   
   	SmartTags("SDC\DB_SDC_ERROR_STAT\_Byte_DB_SDC_ERROR_STAT.F_STAT[XX1].EMS_TS_STAT_VAL.PROFIL") =  			  2 + Eintrag_0 * Laenge_FAULT - Laenge_FAULT + Allg_Offset
   	SmartTags("SDC\DB_SDC_ERROR_STAT\_Byte_DB_SDC_ERROR_STAT.F_STAT[XX2].EMS_TS_STAT_VAL.PROFIL") =  			  2 + Eintrag_1 * Laenge_FAULT - Laenge_FAULT + Allg_Offset
   	SmartTags("SDC\DB_SDC_ERROR_STAT\_Byte_DB_SDC_ERROR_STAT.F_STAT[XX3].EMS_TS_STAT_VAL.PROFIL") =  			  2 + Eintrag_2 * Laenge_FAULT - Laenge_FAULT + Allg_Offset
   	SmartTags("SDC\DB_SDC_ERROR_STAT\_Byte_DB_SDC_ERROR_STAT.F_STAT[XX4].EMS_TS_STAT_VAL.PROFIL") =  			  2 + Eintrag_3 * Laenge_FAULT - Laenge_FAULT + Allg_Offset
   	SmartTags("SDC\DB_SDC_ERROR_STAT\_Byte_DB_SDC_ERROR_STAT.F_STAT[XX5].EMS_TS_STAT_VAL.PROFIL") =  			  2 + Eintrag_4 * Laenge_FAULT - Laenge_FAULT + Allg_Offset
   	SmartTags("SDC\DB_SDC_ERROR_STAT\_Byte_DB_SDC_ERROR_STAT.F_STAT[XX6].EMS_TS_STAT_VAL.PROFIL") =  			  2 + Eintrag_5 * Laenge_FAULT - Laenge_FAULT + Allg_Offset
   	SmartTags("SDC\DB_SDC_ERROR_STAT\_Byte_DB_SDC_ERROR_STAT.F_STAT[XX7].EMS_TS_STAT_VAL.PROFIL") =  			  2 + Eintrag_6 * Laenge_FAULT - Laenge_FAULT + Allg_Offset
   	SmartTags("SDC\DB_SDC_ERROR_STAT\_Byte_DB_SDC_ERROR_STAT.F_STAT[XX8].EMS_TS_STAT_VAL.PROFIL") =  			  2 + Eintrag_7 * Laenge_FAULT - Laenge_FAULT + Allg_Offset
   	SmartTags("SDC\DB_SDC_ERROR_STAT\_Byte_DB_SDC_ERROR_STAT.F_STAT[XX9].EMS_TS_STAT_VAL.PROFIL") =  			  2 + Eintrag_8 * Laenge_FAULT - Laenge_FAULT + Allg_Offset
   	SmartTags("SDC\DB_SDC_ERROR_STAT\_Byte_DB_SDC_ERROR_STAT.F_STAT[X10].EMS_TS_STAT_VAL.PROFIL") =  			  2 + Eintrag_9 * Laenge_FAULT - Laenge_FAULT + Allg_Offset
   
   	SmartTags("SDC\DB_SDC_ERROR_STAT\_Byte_DB_SDC_ERROR_STAT.F_STAT[XX1].EMS_TS_STAT_VAL.DRIVE_POS") =   		  4 + Eintrag_0 * Laenge_FAULT - Laenge_FAULT + Allg_Offset
   	SmartTags("SDC\DB_SDC_ERROR_STAT\_Byte_DB_SDC_ERROR_STAT.F_STAT[XX2].EMS_TS_STAT_VAL.DRIVE_POS") =   		  4 + Eintrag_1 * Laenge_FAULT - Laenge_FAULT + Allg_Offset
   	SmartTags("SDC\DB_SDC_ERROR_STAT\_Byte_DB_SDC_ERROR_STAT.F_STAT[XX3].EMS_TS_STAT_VAL.DRIVE_POS") =   		  4 + Eintrag_2 * Laenge_FAULT - Laenge_FAULT + Allg_Offset
   	SmartTags("SDC\DB_SDC_ERROR_STAT\_Byte_DB_SDC_ERROR_STAT.F_STAT[XX4].EMS_TS_STAT_VAL.DRIVE_POS") =   		  4 + Eintrag_3 * Laenge_FAULT - Laenge_FAULT + Allg_Offset
   	SmartTags("SDC\DB_SDC_ERROR_STAT\_Byte_DB_SDC_ERROR_STAT.F_STAT[XX5].EMS_TS_STAT_VAL.DRIVE_POS") =   		  4 + Eintrag_4 * Laenge_FAULT - Laenge_FAULT + Allg_Offset
   	SmartTags("SDC\DB_SDC_ERROR_STAT\_Byte_DB_SDC_ERROR_STAT.F_STAT[XX6].EMS_TS_STAT_VAL.DRIVE_POS") =   		  4 + Eintrag_5 * Laenge_FAULT - Laenge_FAULT + Allg_Offset
   	SmartTags("SDC\DB_SDC_ERROR_STAT\_Byte_DB_SDC_ERROR_STAT.F_STAT[XX7].EMS_TS_STAT_VAL.DRIVE_POS") =   		  4 + Eintrag_6 * Laenge_FAULT - Laenge_FAULT + Allg_Offset
   	SmartTags("SDC\DB_SDC_ERROR_STAT\_Byte_DB_SDC_ERROR_STAT.F_STAT[XX8].EMS_TS_STAT_VAL.DRIVE_POS") =   		  4 + Eintrag_7 * Laenge_FAULT - Laenge_FAULT + Allg_Offset
   	SmartTags("SDC\DB_SDC_ERROR_STAT\_Byte_DB_SDC_ERROR_STAT.F_STAT[XX9].EMS_TS_STAT_VAL.DRIVE_POS") =   		  4 + Eintrag_8 * Laenge_FAULT - Laenge_FAULT + Allg_Offset
   	SmartTags("SDC\DB_SDC_ERROR_STAT\_Byte_DB_SDC_ERROR_STAT.F_STAT[X10].EMS_TS_STAT_VAL.DRIVE_POS") =   		  4 + Eintrag_9 * Laenge_FAULT - Laenge_FAULT + Allg_Offset
   	
   	SmartTags("SDC\DB_SDC_ERROR_STAT\_Byte_DB_SDC_ERROR_STAT.F_STAT[XX1].EMS_TS_STAT_VAL.HOIST_POS") =   		  8 + Eintrag_0 * Laenge_FAULT - Laenge_FAULT + Allg_Offset
   	SmartTags("SDC\DB_SDC_ERROR_STAT\_Byte_DB_SDC_ERROR_STAT.F_STAT[XX2].EMS_TS_STAT_VAL.HOIST_POS") =   		  8 + Eintrag_1 * Laenge_FAULT - Laenge_FAULT + Allg_Offset
   	SmartTags("SDC\DB_SDC_ERROR_STAT\_Byte_DB_SDC_ERROR_STAT.F_STAT[XX3].EMS_TS_STAT_VAL.HOIST_POS") =   		  8 + Eintrag_2 * Laenge_FAULT - Laenge_FAULT + Allg_Offset
   	SmartTags("SDC\DB_SDC_ERROR_STAT\_Byte_DB_SDC_ERROR_STAT.F_STAT[XX4].EMS_TS_STAT_VAL.HOIST_POS") =   		  8 + Eintrag_3 * Laenge_FAULT - Laenge_FAULT + Allg_Offset
   	SmartTags("SDC\DB_SDC_ERROR_STAT\_Byte_DB_SDC_ERROR_STAT.F_STAT[XX5].EMS_TS_STAT_VAL.HOIST_POS") =   		  8 + Eintrag_4 * Laenge_FAULT - Laenge_FAULT + Allg_Offset
   	SmartTags("SDC\DB_SDC_ERROR_STAT\_Byte_DB_SDC_ERROR_STAT.F_STAT[XX6].EMS_TS_STAT_VAL.HOIST_POS") =   		  8 + Eintrag_5 * Laenge_FAULT - Laenge_FAULT + Allg_Offset
   	SmartTags("SDC\DB_SDC_ERROR_STAT\_Byte_DB_SDC_ERROR_STAT.F_STAT[XX7].EMS_TS_STAT_VAL.HOIST_POS") =   		  8 + Eintrag_6 * Laenge_FAULT - Laenge_FAULT + Allg_Offset
   	SmartTags("SDC\DB_SDC_ERROR_STAT\_Byte_DB_SDC_ERROR_STAT.F_STAT[XX8].EMS_TS_STAT_VAL.HOIST_POS") =   		  8 + Eintrag_7 * Laenge_FAULT - Laenge_FAULT + Allg_Offset
   	SmartTags("SDC\DB_SDC_ERROR_STAT\_Byte_DB_SDC_ERROR_STAT.F_STAT[XX9].EMS_TS_STAT_VAL.HOIST_POS") =   		  8 + Eintrag_8 * Laenge_FAULT - Laenge_FAULT + Allg_Offset
   	SmartTags("SDC\DB_SDC_ERROR_STAT\_Byte_DB_SDC_ERROR_STAT.F_STAT[X10].EMS_TS_STAT_VAL.HOIST_POS") =   		  8 + Eintrag_9 * Laenge_FAULT - Laenge_FAULT + Allg_Offset
   	
   '	SmartTags("SDC\DB_SDC_ERROR_STAT\_Byte_DB_SDC_ERROR_STAT.F_STAT[XX1].EMS_TS_STAT_VAL.TILT_POS")  =   		 10 + Eintrag_0 * Laenge_FAULT - Laenge_FAULT + Allg_Offset
   '	SmartTags("SDC\DB_SDC_ERROR_STAT\_Byte_DB_SDC_ERROR_STAT.F_STAT[XX2].EMS_TS_STAT_VAL.TILT_POS")  =   		 10 + Eintrag_1 * Laenge_FAULT - Laenge_FAULT + Allg_Offset
   '	SmartTags("SDC\DB_SDC_ERROR_STAT\_Byte_DB_SDC_ERROR_STAT.F_STAT[XX3].EMS_TS_STAT_VAL.TILT_POS")  =   		 10 + Eintrag_2 * Laenge_FAULT - Laenge_FAULT + Allg_Offset
   '	SmartTags("SDC\DB_SDC_ERROR_STAT\_Byte_DB_SDC_ERROR_STAT.F_STAT[XX4].EMS_TS_STAT_VAL.TILT_POS")  =   		 10 + Eintrag_3 * Laenge_FAULT - Laenge_FAULT + Allg_Offset
   '	SmartTags("SDC\DB_SDC_ERROR_STAT\_Byte_DB_SDC_ERROR_STAT.F_STAT[XX5].EMS_TS_STAT_VAL.TILT_POS")  =   		 10 + Eintrag_4 * Laenge_FAULT - Laenge_FAULT + Allg_Offset
   '	SmartTags("SDC\DB_SDC_ERROR_STAT\_Byte_DB_SDC_ERROR_STAT.F_STAT[XX6].EMS_TS_STAT_VAL.TILT_POS")  =   		 10 + Eintrag_5 * Laenge_FAULT - Laenge_FAULT + Allg_Offset
   '	SmartTags("SDC\DB_SDC_ERROR_STAT\_Byte_DB_SDC_ERROR_STAT.F_STAT[XX7].EMS_TS_STAT_VAL.TILT_POS")  =   		 10 + Eintrag_6 * Laenge_FAULT - Laenge_FAULT + Allg_Offset
   '	SmartTags("SDC\DB_SDC_ERROR_STAT\_Byte_DB_SDC_ERROR_STAT.F_STAT[XX8].EMS_TS_STAT_VAL.TILT_POS")  =   		 10 + Eintrag_7 * Laenge_FAULT - Laenge_FAULT + Allg_Offset
   '	SmartTags("SDC\DB_SDC_ERROR_STAT\_Byte_DB_SDC_ERROR_STAT.F_STAT[XX9].EMS_TS_STAT_VAL.TILT_POS")  =   		 10 + Eintrag_8 * Laenge_FAULT - Laenge_FAULT + Allg_Offset
   '	SmartTags("SDC\DB_SDC_ERROR_STAT\_Byte_DB_SDC_ERROR_STAT.F_STAT[X10].EMS_TS_STAT_VAL.TILT_POS")  =   		 10 + Eintrag_9 * Laenge_FAULT - Laenge_FAULT + Allg_Offset
   	
   	SmartTags("SDC\DB_SDC_ERROR_STAT\_Byte_DB_SDC_ERROR_STAT.F_STAT[XX1].EMS_TS_STAT_VAL.ERROR")  	 =   		 10 + Eintrag_0 * Laenge_FAULT - Laenge_FAULT + Allg_Offset
   	SmartTags("SDC\DB_SDC_ERROR_STAT\_Byte_DB_SDC_ERROR_STAT.F_STAT[XX2].EMS_TS_STAT_VAL.ERROR")  	 =   		 10 + Eintrag_1 * Laenge_FAULT - Laenge_FAULT + Allg_Offset
   	SmartTags("SDC\DB_SDC_ERROR_STAT\_Byte_DB_SDC_ERROR_STAT.F_STAT[XX3].EMS_TS_STAT_VAL.ERROR")  	 =   		 10 + Eintrag_2 * Laenge_FAULT - Laenge_FAULT + Allg_Offset
   	SmartTags("SDC\DB_SDC_ERROR_STAT\_Byte_DB_SDC_ERROR_STAT.F_STAT[XX4].EMS_TS_STAT_VAL.ERROR")  	 =   		 10 + Eintrag_3 * Laenge_FAULT - Laenge_FAULT + Allg_Offset
   	SmartTags("SDC\DB_SDC_ERROR_STAT\_Byte_DB_SDC_ERROR_STAT.F_STAT[XX5].EMS_TS_STAT_VAL.ERROR")  	 =   		 10 + Eintrag_4 * Laenge_FAULT - Laenge_FAULT + Allg_Offset
   	SmartTags("SDC\DB_SDC_ERROR_STAT\_Byte_DB_SDC_ERROR_STAT.F_STAT[XX6].EMS_TS_STAT_VAL.ERROR")  	 =   		 10 + Eintrag_5 * Laenge_FAULT - Laenge_FAULT + Allg_Offset
   	SmartTags("SDC\DB_SDC_ERROR_STAT\_Byte_DB_SDC_ERROR_STAT.F_STAT[XX7].EMS_TS_STAT_VAL.ERROR")  	 =   		 10 + Eintrag_6 * Laenge_FAULT - Laenge_FAULT + Allg_Offset
   	SmartTags("SDC\DB_SDC_ERROR_STAT\_Byte_DB_SDC_ERROR_STAT.F_STAT[XX8].EMS_TS_STAT_VAL.ERROR")  	 =   		 10 + Eintrag_7 * Laenge_FAULT - Laenge_FAULT + Allg_Offset
   	SmartTags("SDC\DB_SDC_ERROR_STAT\_Byte_DB_SDC_ERROR_STAT.F_STAT[XX9].EMS_TS_STAT_VAL.ERROR")  	 =   		 10 + Eintrag_8 * Laenge_FAULT - Laenge_FAULT + Allg_Offset
   	SmartTags("SDC\DB_SDC_ERROR_STAT\_Byte_DB_SDC_ERROR_STAT.F_STAT[X10].EMS_TS_STAT_VAL.ERROR")  	 =   		 10 + Eintrag_9 * Laenge_FAULT - Laenge_FAULT + Allg_Offset
   
   	SmartTags("SDC\DB_SDC_ERROR_STAT\_Byte_DB_SDC_ERROR_STAT.F_STAT[XX1].EMS_TS_STAT_VAL.DRIVE_POS_PERC") =   	 12 + Eintrag_0 * Laenge_FAULT - Laenge_FAULT + Allg_Offset
   	SmartTags("SDC\DB_SDC_ERROR_STAT\_Byte_DB_SDC_ERROR_STAT.F_STAT[XX2].EMS_TS_STAT_VAL.DRIVE_POS_PERC") =   	 12 + Eintrag_1 * Laenge_FAULT - Laenge_FAULT + Allg_Offset
   	SmartTags("SDC\DB_SDC_ERROR_STAT\_Byte_DB_SDC_ERROR_STAT.F_STAT[XX3].EMS_TS_STAT_VAL.DRIVE_POS_PERC") =   	 12 + Eintrag_2 * Laenge_FAULT - Laenge_FAULT + Allg_Offset
   	SmartTags("SDC\DB_SDC_ERROR_STAT\_Byte_DB_SDC_ERROR_STAT.F_STAT[XX4].EMS_TS_STAT_VAL.DRIVE_POS_PERC") =   	 12 + Eintrag_3 * Laenge_FAULT - Laenge_FAULT + Allg_Offset
   	SmartTags("SDC\DB_SDC_ERROR_STAT\_Byte_DB_SDC_ERROR_STAT.F_STAT[XX5].EMS_TS_STAT_VAL.DRIVE_POS_PERC") =   	 12 + Eintrag_4 * Laenge_FAULT - Laenge_FAULT + Allg_Offset
   	SmartTags("SDC\DB_SDC_ERROR_STAT\_Byte_DB_SDC_ERROR_STAT.F_STAT[XX6].EMS_TS_STAT_VAL.DRIVE_POS_PERC") =   	 12 + Eintrag_5 * Laenge_FAULT - Laenge_FAULT + Allg_Offset
   	SmartTags("SDC\DB_SDC_ERROR_STAT\_Byte_DB_SDC_ERROR_STAT.F_STAT[XX7].EMS_TS_STAT_VAL.DRIVE_POS_PERC") =   	 12 + Eintrag_6 * Laenge_FAULT - Laenge_FAULT + Allg_Offset
   	SmartTags("SDC\DB_SDC_ERROR_STAT\_Byte_DB_SDC_ERROR_STAT.F_STAT[XX8].EMS_TS_STAT_VAL.DRIVE_POS_PERC") =   	 12 + Eintrag_7 * Laenge_FAULT - Laenge_FAULT + Allg_Offset
   	SmartTags("SDC\DB_SDC_ERROR_STAT\_Byte_DB_SDC_ERROR_STAT.F_STAT[XX9].EMS_TS_STAT_VAL.DRIVE_POS_PERC") =   	 12 + Eintrag_8 * Laenge_FAULT - Laenge_FAULT + Allg_Offset
   	SmartTags("SDC\DB_SDC_ERROR_STAT\_Byte_DB_SDC_ERROR_STAT.F_STAT[X10].EMS_TS_STAT_VAL.DRIVE_POS_PERC") =   	 12 + Eintrag_9 * Laenge_FAULT - Laenge_FAULT + Allg_Offset
   	
   	SmartTags("SDC\DB_SDC_ERROR_STAT\_Byte_DB_SDC_ERROR_STAT.F_STAT[XX1].EMS_TS_STAT_VAL.SEK") 			=   	 14 + Eintrag_0 * Laenge_FAULT - Laenge_FAULT + Allg_Offset
   	SmartTags("SDC\DB_SDC_ERROR_STAT\_Byte_DB_SDC_ERROR_STAT.F_STAT[XX2].EMS_TS_STAT_VAL.SEK") 			=   	 14 + Eintrag_1 * Laenge_FAULT - Laenge_FAULT + Allg_Offset
   	SmartTags("SDC\DB_SDC_ERROR_STAT\_Byte_DB_SDC_ERROR_STAT.F_STAT[XX3].EMS_TS_STAT_VAL.SEK") 			=   	 14 + Eintrag_2 * Laenge_FAULT - Laenge_FAULT + Allg_Offset
   	SmartTags("SDC\DB_SDC_ERROR_STAT\_Byte_DB_SDC_ERROR_STAT.F_STAT[XX4].EMS_TS_STAT_VAL.SEK") 			=   	 14 + Eintrag_3 * Laenge_FAULT - Laenge_FAULT + Allg_Offset
   	SmartTags("SDC\DB_SDC_ERROR_STAT\_Byte_DB_SDC_ERROR_STAT.F_STAT[XX5].EMS_TS_STAT_VAL.SEK") 			=   	 14 + Eintrag_4 * Laenge_FAULT - Laenge_FAULT + Allg_Offset
   	SmartTags("SDC\DB_SDC_ERROR_STAT\_Byte_DB_SDC_ERROR_STAT.F_STAT[XX6].EMS_TS_STAT_VAL.SEK") 			=   	 14 + Eintrag_5 * Laenge_FAULT - Laenge_FAULT + Allg_Offset
   	SmartTags("SDC\DB_SDC_ERROR_STAT\_Byte_DB_SDC_ERROR_STAT.F_STAT[XX7].EMS_TS_STAT_VAL.SEK") 			=   	 14 + Eintrag_6 * Laenge_FAULT - Laenge_FAULT + Allg_Offset
   	SmartTags("SDC\DB_SDC_ERROR_STAT\_Byte_DB_SDC_ERROR_STAT.F_STAT[XX8].EMS_TS_STAT_VAL.SEK") 			=   	 14 + Eintrag_7 * Laenge_FAULT - Laenge_FAULT + Allg_Offset
   	SmartTags("SDC\DB_SDC_ERROR_STAT\_Byte_DB_SDC_ERROR_STAT.F_STAT[XX9].EMS_TS_STAT_VAL.SEK") 			=   	 14 + Eintrag_8 * Laenge_FAULT - Laenge_FAULT + Allg_Offset
   	SmartTags("SDC\DB_SDC_ERROR_STAT\_Byte_DB_SDC_ERROR_STAT.F_STAT[X10].EMS_TS_STAT_VAL.SEK") 			=   	 14 + Eintrag_9 * Laenge_FAULT - Laenge_FAULT + Allg_Offset
   	
   	SmartTags("SDC\DB_SDC_ERROR_STAT\_Byte_DB_SDC_ERROR_STAT.F_STAT[XX1].F") = 									 16 + Eintrag_0 * Laenge_FAULT - Laenge_FAULT + Allg_Offset
   	SmartTags("SDC\DB_SDC_ERROR_STAT\_Byte_DB_SDC_ERROR_STAT.F_STAT[XX2].F") = 									 16 + Eintrag_1 * Laenge_FAULT - Laenge_FAULT + Allg_Offset
   	SmartTags("SDC\DB_SDC_ERROR_STAT\_Byte_DB_SDC_ERROR_STAT.F_STAT[XX3].F") = 									 16 + Eintrag_2 * Laenge_FAULT - Laenge_FAULT + Allg_Offset
   	SmartTags("SDC\DB_SDC_ERROR_STAT\_Byte_DB_SDC_ERROR_STAT.F_STAT[XX4].F") = 									 16 + Eintrag_3 * Laenge_FAULT - Laenge_FAULT + Allg_Offset
   	SmartTags("SDC\DB_SDC_ERROR_STAT\_Byte_DB_SDC_ERROR_STAT.F_STAT[XX5].F") = 									 16 + Eintrag_4 * Laenge_FAULT - Laenge_FAULT + Allg_Offset
   	SmartTags("SDC\DB_SDC_ERROR_STAT\_Byte_DB_SDC_ERROR_STAT.F_STAT[XX6].F") = 									 16 + Eintrag_5 * Laenge_FAULT - Laenge_FAULT + Allg_Offset
   	SmartTags("SDC\DB_SDC_ERROR_STAT\_Byte_DB_SDC_ERROR_STAT.F_STAT[XX7].F") = 									 16 + Eintrag_6 * Laenge_FAULT - Laenge_FAULT + Allg_Offset
   	SmartTags("SDC\DB_SDC_ERROR_STAT\_Byte_DB_SDC_ERROR_STAT.F_STAT[XX8].F") = 									 16 + Eintrag_7 * Laenge_FAULT - Laenge_FAULT + Allg_Offset
   	SmartTags("SDC\DB_SDC_ERROR_STAT\_Byte_DB_SDC_ERROR_STAT.F_STAT[XX9].F") = 									 16 + Eintrag_8 * Laenge_FAULT - Laenge_FAULT + Allg_Offset
   	SmartTags("SDC\DB_SDC_ERROR_STAT\_Byte_DB_SDC_ERROR_STAT.F_STAT[X10].F") = 									 16 + Eintrag_9 * Laenge_FAULT - Laenge_FAULT + Allg_Offset
   	
   	SmartTags("SDC\DB_SDC_ERROR_STAT\_Byte_DB_SDC_ERROR_STAT.F_STAT[XX1].F_DATE") = 							 20 + Eintrag_0 * Laenge_FAULT - Laenge_FAULT + Allg_Offset
   	SmartTags("SDC\DB_SDC_ERROR_STAT\_Byte_DB_SDC_ERROR_STAT.F_STAT[XX2].F_DATE") = 							 20 + Eintrag_1 * Laenge_FAULT - Laenge_FAULT + Allg_Offset
   	SmartTags("SDC\DB_SDC_ERROR_STAT\_Byte_DB_SDC_ERROR_STAT.F_STAT[XX3].F_DATE") = 							 20 + Eintrag_2 * Laenge_FAULT - Laenge_FAULT + Allg_Offset
   	SmartTags("SDC\DB_SDC_ERROR_STAT\_Byte_DB_SDC_ERROR_STAT.F_STAT[XX4].F_DATE") = 							 20 + Eintrag_3 * Laenge_FAULT - Laenge_FAULT + Allg_Offset
   	SmartTags("SDC\DB_SDC_ERROR_STAT\_Byte_DB_SDC_ERROR_STAT.F_STAT[XX5].F_DATE") = 							 20 + Eintrag_4 * Laenge_FAULT - Laenge_FAULT + Allg_Offset
   	SmartTags("SDC\DB_SDC_ERROR_STAT\_Byte_DB_SDC_ERROR_STAT.F_STAT[XX6].F_DATE") = 							 20 + Eintrag_5 * Laenge_FAULT - Laenge_FAULT + Allg_Offset
   	SmartTags("SDC\DB_SDC_ERROR_STAT\_Byte_DB_SDC_ERROR_STAT.F_STAT[XX7].F_DATE") = 							 20 + Eintrag_6 * Laenge_FAULT - Laenge_FAULT + Allg_Offset
   	SmartTags("SDC\DB_SDC_ERROR_STAT\_Byte_DB_SDC_ERROR_STAT.F_STAT[XX8].F_DATE") = 							 20 + Eintrag_7 * Laenge_FAULT - Laenge_FAULT + Allg_Offset
   	SmartTags("SDC\DB_SDC_ERROR_STAT\_Byte_DB_SDC_ERROR_STAT.F_STAT[XX9].F_DATE") = 							 20 + Eintrag_8 * Laenge_FAULT - Laenge_FAULT + Allg_Offset
   	SmartTags("SDC\DB_SDC_ERROR_STAT\_Byte_DB_SDC_ERROR_STAT.F_STAT[X10].F_DATE") = 							 20 + Eintrag_9 * Laenge_FAULT - Laenge_FAULT + Allg_Offset
   	
   	
   	
   	

VB script "SDC_ERRORS"
   'HINWEIS:
   ' Beim Erstellen von Skripten können Sie mit <Strg+Leertaste> vordefinierte 
   ' Systemfunktionen in das neue Skript einbinden.
   ' Das HMIRuntime-Objekt ermöglicht einfachen Zugriff auf die Objekte des
   ' WinCC flexible Objektmodells, ihre Methoden und ihre Eigenschaften.
   ' Für ein komfortables Auswählen einer Objektreferenz betätigen Sie bitte <Alt+Rechts>.
   ' Komplexe Skripte können Sie mit Sprachelementen der Programmiersprache
   ' VBScript erstellen.
   ' Der Zugriff auf WinCC flexible Variablen erfolgt direkt über den Variablennamen,
   ' z.B. Tag = 5
   
   '________________________________________________________________________________
   '
   
   ' Groiß Andreas
   ' Siemens AG Österreich 
   ' Linz Kraußstraße 1-7 
   ' RC-AT I-IA AS-FA-SO-AE2
   ' 07.07.2015
   Dim EMS_Nr ' EMS Number
   Dim Laenge_Errors ' Länge Errors
   Dim Allg_Offset ' Allg Offset
   Dim OffsetEMS_Errors ' Offset je EMS von Errors
   
   
   ' INIT-------------------------------------------------------------
   EMS_Nr = EMS_Nr_IN
   
   If (EMS_Nr_IN < SmartTags("DB_SDC_ERRORS_HEADER.MIN_NR_EMS")) Or (EMS_Nr_IN > SmartTags("DB_SDC_ERRORS_HEADER.MAX_NR_EMS")) Then
   	EMS_Nr = SmartTags("DB_SDC_ERRORS_HEADER.MIN_NR_EMS")
   End If	
   
   If EMS_Nr_IN < 1 Then
   	EMS_Nr = 1
   End If	
   
   
   '##############################################
   ' VISU Sucht sich Sektions daten:
   '##############################################
   Laenge_Errors = SmartTags("DB_SDC_ERRORS_HEADER.LAENGE_EMS_StörungS")
   
   Allg_Offset = SmartTags("DB_SDC_ERRORS_HEADER.START_EMS")
   
   OffsetEMS_Errors = EMS_Nr * Laenge_Errors - Laenge_Errors + Allg_Offset
   
   SmartTags("_Byte_DB_SDC_ERRORS.EMS[XXX].GEN_1") =						  0 + OffsetEMS_Errors
   SmartTags("_Byte_DB_SDC_ERRORS.EMS[XXX].GEN_2") =						  2 + OffsetEMS_Errors
   SmartTags("_Byte_DB_SDC_ERRORS.EMS[XXX].GEN_3") =						  4 + OffsetEMS_Errors
   SmartTags("_Byte_DB_SDC_ERRORS.EMS[XXX].GEN_4") =						  6 + OffsetEMS_Errors
   
   SmartTags("_Byte_DB_SDC_ERRORS.EMS[XXX].DRIVE_1") =						  8 + OffsetEMS_Errors
   SmartTags("_Byte_DB_SDC_ERRORS.EMS[XXX].DRIVE_2") =						 10 + OffsetEMS_Errors
   SmartTags("_Byte_DB_SDC_ERRORS.EMS[XXX].FC_DRIVE_1") =					 12 + OffsetEMS_Errors
   SmartTags("_Byte_DB_SDC_ERRORS.EMS[XXX].SAFETY_DRIVE") =				 14 + OffsetEMS_Errors
   SmartTags("_Byte_DB_SDC_ERRORS.EMS[XXX].FC_DRIVE_2") =					 16 + OffsetEMS_Errors
   
   SmartTags("_Byte_DB_SDC_ERRORS.EMS[XXX].HOIST_1") =						 18 + OffsetEMS_Errors
   SmartTags("_Byte_DB_SDC_ERRORS.EMS[XXX].HOIST_2") =						 20 + OffsetEMS_Errors
   SmartTags("_Byte_DB_SDC_ERRORS.EMS[XXX].FC_HOIST_1") =					 22 + OffsetEMS_Errors
   SmartTags("_Byte_DB_SDC_ERRORS.EMS[XXX].SAFETY_HOIST") =				 24 + OffsetEMS_Errors
   SmartTags("_Byte_DB_SDC_ERRORS.EMS[XXX].FC_HOIST_2") =					 26 + OffsetEMS_Errors
   
   'SmartTags("_Byte_DB_SDC_ERRORS.EMS[XXX].TILT_1") =						 28 + OffsetEMS_Errors
   'SmartTags("_Byte_DB_SDC_ERRORS.EMS[XXX].TILT_2") =						 30 + OffsetEMS_Errors
   'SmartTags("_Byte_DB_SDC_ERRORS.EMS[XXX].FC_TILT_1") =					 32 + OffsetEMS_Errors
   'SmartTags("_Byte_DB_SDC_ERRORS.EMS[XXX].SAFETY_TILT") =		     		 34 + OffsetEMS_Errors
   'SmartTags("_Byte_DB_SDC_ERRORS.EMS[XXX].FC_TILT_2") =					 36 + OffsetEMS_Errors
   
   SmartTags("_Byte_DB_SDC_ERRORS.EMS[XXX].SDC") =	    					 48 + OffsetEMS_Errors

VB script "SDC_GLOBAL_REFERENCE_PROFIL"
   'HINWEIS:
   ' Beim Erstellen von Skripten können Sie mit <Strg+Leertaste> vordefinierte 
   ' Systemfunktionen in das neue Skript einbinden.
   ' Das HMIRuntime-Objekt ermöglicht einfachen Zugriff auf die Objekte des
   ' WinCC flexible Objektmodells, ihre Methoden und ihre Eigenschaften.
   ' Für ein komfortables Auswählen einer Objektreferenz betätigen Sie bitte <Alt+Rechts>.
   ' Komplexe Skripte können Sie mit Sprachelementen der Programmiersprache
   ' VBScript erstellen.
   ' Der Zugriff auf WinCC flexible Variablen erfolgt direkt über den Variablennamen,
   ' z.B. Tag = 5
   
   '________________________________________________________________________________
   '
   
   ' Groiß Andreas
   ' Siemens AG Österreich 
   ' Linz Kraußstraße 1-7 
   ' RC-AT I-IA AS-FA-SO-AE2
   ' 02.08.2013
   
   
   'Profil Referenz
   
   Dim Profil_Nr ' Sektion Number
   Dim Laenge_Profil ' Länge Profil
   Dim Profil_Offset ' Allg Profil Offset
   
   'Profilnummer - 1 da 2 Profile angezeigt werden
   If SmartTags("DB_SDC_GLOBAL_REFERENCE_HEADER.MIN_PROFIL") <= Profil_Nr_IN And (SmartTags("DB_SDC_GLOBAL_REFERENCE_HEADER.MAX_PROFIL") - 1) >= Profil_Nr_IN Then
    Profil_Nr = Profil_Nr_IN
   Else
    Profil_Nr = "SDC\DB_SDC_GLOBAL_REFERENCE\DB_SDC_GLOBAL_REFERENCE.HEADER.MIN_PROFIL"	 
   End If	 
   
   Laenge_Profil = SmartTags("DB_SDC_GLOBAL_REFERENCE_HEADER.LAENGE_PROFIL")
   Profil_Offset = SmartTags("DB_SDC_GLOBAL_REFERENCE_HEADER.START_PROFIL")
   
     SmartTags("_DB_SDC_GLOBAL_REFERENCE.PROFIL[XX].SORTE_Byte") = Profil_Nr * Laenge_Profil - Laenge_Profil + Profil_Offset 
     SmartTags("_DB_SDC_GLOBAL_REFERENCE.PROFIL[XX+1].SORTE_Byte") = (Profil_Nr +1) * Laenge_Profil - Laenge_Profil + Profil_Offset 

VB script "SDC_PN"
   If SmartTags("_intern_BILD_Nr")= 100 Or SmartTags("_intern_BILD_Nr")= 101 Then
   	If SmartTags("PN_PB\PN\IOSys_ID") = 100 Then
         Call b431313b-d6b5-4a28-b630-23a386ef7180(PN_100, SmartTags("PN_PB\PN\Teiln_Nr")+1, Null)
   	End If
   	If SmartTags("PN_PB\PN\IOSys_ID") = 101 Then
         Call b431313b-d6b5-4a28-b630-23a386ef7180(PN_101, SmartTags("PN_PB\PN\Teiln_Nr")+1, Null)
   	End If 
   End If

VB script "SDC_TS_IF"
   'HINWEIS:
   ' Beim Erstellen von Skripten können Sie mit <Strg+Leertaste> vordefinierte 
   ' Systemfunktionen in das neue Skript einbinden.
   ' Das HMIRuntime-Objekt ermöglicht einfachen Zugriff auf die Objekte des
   ' WinCC flexible Objektmodells, ihre Methoden und ihre Eigenschaften.
   ' Für ein komfortables Auswählen einer Objektreferenz betätigen Sie bitte <Alt+Rechts>.
   ' Komplexe Skripte können Sie mit Sprachelementen der Programmiersprache
   ' VBScript erstellen.
   ' Der Zugriff auf WinCC flexible Variablen erfolgt direkt über den Variablennamen,
   ' z.B. Tag = 5
   
   '________________________________________________________________________________
   '
   
   ' Groiß Andreas
   ' Siemens AG Österreich 
   ' Linz Kraußstraße 1-7 
   ' RC-AT I-IA AS-FA-SO-AE2
   ' 07.07.2015
   Dim TS_Nr ' Sektion Number
   Dim Laenge_Data ' Länge TS
   Dim Allg_Offset ' Allg TS Offset
   Dim OffsetTS ' TS Offset
   Dim OffsetSTAT ' TS Stat Offset
   Dim HMISekDaten_Offset ' HMI Sektionsdaten Offset
   Dim HMI_Nr ' HMI Nummer
   
   '##############################################
   ' S7 sucht sich Sektionsdaten:
   '##############################################
   
   ' INIT-------------------------------------------------------------
   SmartTags("_DB_SDC_TS_IF_COMMAND.HEADER.DB_NR") = SmartTags("DB_SDC_TS_IF_HMI_HEADER.DB_NR")
   SmartTags("_DB_SDC_TS_IF_STATUS.HEADER.DB_NR") = SmartTags("DB_SDC_TS_IF_HMI_HEADER.DB_NR")
   
   If (SmartTags("SDC\_TS_Nr") < SmartTags("DB_SDC_GLOBAL_SEK_MIN")) Or (SmartTags("SDC\_TS_Nr") > SmartTags("DB_SDC_GLOBAL_SEK_MAX")) Then
   	SmartTags("SDC\_TS_Nr") = 	SmartTags("DB_SDC_GLOBAL_SEK_MIN")
   End If	
   
   If (SmartTags("SDC\_TS_Nr") < 1) Then
   	SmartTags("SDC\_TS_Nr") = 1
   End If	
   
   HMISekDaten_Offset = SmartTags("DB_SDC_TS_IF_HMI_HEADER.OFFEST_HMI_DATA")
   HMI_Nr = SmartTags("_intern_Pult_Nr")
   
   Laenge_Data = SmartTags("DB_SDC_TS_IF_HMI_HEADER.LAENGE_SEK_COM") + SmartTags("DB_SDC_TS_IF_HMI_HEADER.LAENGE_SEK_STAT")
   
   Allg_Offset = SmartTags("DB_SDC_TS_IF_HMI_HEADER.START_HMI")
      
   OffsetTS = HMI_Nr * (Laenge_Data + HMISekDaten_Offset)  - Laenge_Data + Allg_Offset
   	
      SmartTags("_DB_SDC_TS_IF_HMI.HMI_Byte_00") = 0 + OffsetTS - HMISekDaten_Offset
      SmartTags("_DB_SDC_TS_IF_HMI.HMI_Byte_02") = 2 + OffsetTS - HMISekDaten_Offset	
      SmartTags("_DB_SDC_TS_IF_HMI.HMI_Byte_04") = 4 + OffsetTS - HMISekDaten_Offset	
      SmartTags("_DB_SDC_TS_IF_HMI.HMI_Byte_06") = 6 + OffsetTS - HMISekDaten_Offset	
      SmartTags("_DB_SDC_TS_IF_HMI.HMI_Byte_08") = 8 + OffsetTS - HMISekDaten_Offset	
      SmartTags("_DB_SDC_TS_IF_HMI.HMI_Byte_09") = 9 + OffsetTS - HMISekDaten_Offset	
      SmartTags("_DB_SDC_TS_IF_HMI.HMI_Byte_10") = 10 + OffsetTS - HMISekDaten_Offset	
      SmartTags("_DB_SDC_TS_IF_HMI.HMI_Byte_12") = 12 + OffsetTS - HMISekDaten_Offset		
      SmartTags("_DB_SDC_TS_IF_HMI.HMI_Byte_14") = 14 + OffsetTS - HMISekDaten_Offset	
      SmartTags("_DB_SDC_TS_IF_HMI.HMI_Byte_16") = 16 + OffsetTS - HMISekDaten_Offset	
      SmartTags("_DB_SDC_TS_IF_HMI.HMI_Byte_18") = 18 + OffsetTS - HMISekDaten_Offset	
      SmartTags("_DB_SDC_TS_IF_HMI.HMI_Byte_19") = 19 + OffsetTS - HMISekDaten_Offset
      
   ' COMMAND
   SmartTags("_Byte_DB_SDC_TS_IF_COMMAND.SEK[XXX].VAL.PROFIL") =						  0 + OffsetTS
   SmartTags("_Byte_DB_SDC_TS_IF_COMMAND.SEK[XXX].VAL.D_SETSPEED") =					  2 + OffsetTS
   SmartTags("_Byte_DB_SDC_TS_IF_COMMAND.SEK[XXX].VAL.D_POS_OFFS") =					  6 + OffsetTS
   
   SmartTags("_Byte_DB_SDC_TS_IF_COMMAND.SEK[XXX].BIT1") =					 			 10 + OffsetTS
   SmartTags("_Byte_DB_SDC_TS_IF_COMMAND.SEK[XXX].BIT2") =					 			 12 + OffsetTS
   'SmartTags("_Byte_DB_SDC_TS_IF_COMMAND.SEK[XXX].BIT3") =					 			 12 + OffsetTS
   
   SmartTags("_Byte_DB_SDC_TS_IF_COMMAND.SEK[XXX].FKT_SET") =				 			 14 + OffsetTS
   SmartTags("_Byte_DB_SDC_TS_IF_COMMAND.SEK[XXX].FKT_RESET") =			 			 16 + OffsetTS
   
   ' STATUS
   OffsetSTAT =  SmartTags("DB_SDC_TS_IF_HMI_HEADER.OFFEST_SEK_STAT")
   
   SmartTags("_Byte_DB_SDC_TS_IF_STATUS.SEK[XXX].VAL.EMS_ID") =						  0 + OffsetTS + OffsetSTAT
   SmartTags("_Byte_DB_SDC_TS_IF_STATUS.SEK[XXX].VAL.PROFIL") =						  2 + OffsetTS + OffsetSTAT
   SmartTags("_Byte_DB_SDC_TS_IF_STATUS.SEK[XXX].VAL.DRIVE_POS") =						  4 + OffsetTS + OffsetSTAT
   SmartTags("_Byte_DB_SDC_TS_IF_STATUS.SEK[XXX].VAL.HOIST_POS") =						  8 + OffsetTS + OffsetSTAT
   'SmartTags("_Byte_DB_SDC_TS_IF_STATUS.SEK[XXX].VAL.TILT_POS") =						 10 + OffsetTS + OffsetSTAT
   SmartTags("_Byte_DB_SDC_TS_IF_STATUS.SEK[XXX].VAL.ERROR") =							 10 + OffsetTS + OffsetSTAT
   SmartTags("_Byte_DB_SDC_TS_IF_STATUS.SEK[XXX].VAL.DRIVE_POS_PERC") =				 12 + OffsetTS + OffsetSTAT
   SmartTags("_Byte_DB_SDC_TS_IF_STATUS.SEK[XXX].VAL.SEK") =							 14 + OffsetTS + OffsetSTAT
   
   SmartTags("_Byte_DB_SDC_TS_IF_STATUS.SEK[XXX].BIT1") =					 			 16 + OffsetTS + OffsetSTAT
   SmartTags("_Byte_DB_SDC_TS_IF_STATUS.SEK[XXX].BIT2") =					 			 18 + OffsetTS + OffsetSTAT
   SmartTags("_Byte_DB_SDC_TS_IF_STATUS.SEK[XXX].BIT3") =					 			 20 + OffsetTS + OffsetSTAT
   'SmartTags("_Byte_DB_SDC_TS_IF_STATUS.SEK[XXX].BIT4") =					 			 24 + OffsetTS + OffsetSTAT
   
   SmartTags("_Byte_DB_SDC_TS_IF_STATUS.SEK[XXX].SORTE") =					 			 22 + OffsetTS + OffsetSTAT
   
   SmartTags("_Byte_DB_SDC_TS_IF_STATUS.SEK[XXX].FKT_SET") =				 			 26 + OffsetTS + OffsetSTAT
   
   
   SmartTags("DB_SDC_TS_IF_HMI.HMI[XX].SEK_Nr") = SmartTags("SDC\_TS_Nr")
   
   '##############################################
   ' VISU Sucht sich Sektions daten:
   '##############################################
   
   '################################################
   '################### COMMANDS ###################
   '################################################
   
   ' INIT-------------------------------------------------------------
   'SmartTags("_Byte_DB_SDC_TS_IF_COMMAND.HEADER.DB_NR") = SmartTags("DB_SDC_TS_IF_COMMAND.HEADER.DB_NR")
   
   'If (SmartTags("SDC\_TS_Nr") < SmartTags("DB_SDC_TS_IF_COMMAND.HEADER.SEK_MIN")) Or (SmartTags("SDC\_TS_Nr") > SmartTags("DB_SDC_TS_IF_COMMAND.HEADER.SEK_MAX")) Then
   '	If (SmartTags("SDC\_TS_Nr") < SmartTags("DB_SDC_TS_IF_COMMAND_2.HEADER.SEK_MIN")) Or (SmartTags("SDC\_TS_Nr") > SmartTags("DB_SDC_TS_IF_COMMAND_2.HEADER.SEK_MAX")) Then
   '		SmartTags("SDC\_TS_Nr") = 	SmartTags("DB_SDC_TS_IF_COMMAND.HEADER.SEK_MIN")
   '	End If		
   'End If	
   	
   
   'If (SmartTags("SDC\_TS_Nr") < 1) Then
   '	SmartTags("SDC\_TS_Nr") = 1
   'End If	
   
   'TS_Nr = SmartTags("SDC\_TS_Nr")
   
   'If (SmartTags("SDC\_TS_Nr") >= SmartTags("DB_SDC_TS_IF_COMMAND_2.HEADER.SEK_MIN")) And (SmartTags("SDC\_TS_Nr") <= SmartTags("DB_SDC_TS_IF_COMMAND_2.HEADER.SEK_MAX")) Then
   '	SmartTags("_Byte_DB_SDC_TS_IF_COMMAND.HEADER.DB_NR") = SmartTags("DB_SDC_TS_IF_COMMAND_2.HEADER.DB_NR")	
   '	TS_Nr = SmartTags("SDC\_TS_Nr") - SmartTags("DB_SDC_TS_IF_COMMAND_2.HEADER.SEK_MIN") + 1
   'End If	
   
   
   'Laenge_Data = SmartTags("DB_SDC_TS_IF_COMMAND.HEADER.LAENGE_SEK_DATA")
   
   'Allg_Offset = SmartTags("DB_SDC_TS_IF_COMMAND.HEADER.START_DAT")
   
   'OffsetTS = TS_Nr  * Laenge_Data - Laenge_Data + Allg_Offset
   
   'SmartTags("_Byte_DB_SDC_TS_IF_COMMAND.SEK[XXX].VAL.PROFIL") =						  0 + OffsetTS
   'SmartTags("_Byte_DB_SDC_TS_IF_COMMAND.SEK[XXX].VAL.D_SETSPEED") =					  2 + OffsetTS
   'SmartTags("_Byte_DB_SDC_TS_IF_COMMAND.SEK[XXX].VAL.D_POS_OFFS") =					  6 + OffsetTS
   
   'SmartTags("_Byte_DB_SDC_TS_IF_COMMAND.SEK[XXX].BIT1") =					 			  8 + OffsetTS
   'SmartTags("_Byte_DB_SDC_TS_IF_COMMAND.SEK[XXX].BIT2") =					 			 10 + OffsetTS
   'SmartTags("_Byte_DB_SDC_TS_IF_COMMAND.SEK[XXX].BIT3") =					 			 12 + OffsetTS
   
   'SmartTags("_Byte_DB_SDC_TS_IF_COMMAND.SEK[XXX].FKT_SET") =				 			 14 + OffsetTS
   'SmartTags("_Byte_DB_SDC_TS_IF_COMMAND.SEK[XXX].FKT_RESET") =			 			 16 + OffsetTS
   
   
   '################################################
   '################### STATUS ###################
   '################################################
   
   ' INIT-------------------------------------------------------------
   'SmartTags("_Byte_DB_SDC_TS_IF_STATUS.HEADER.DB_NR") = SmartTags("DB_SDC_TS_IF_STATUS.HEADER.DB_NR")
   
   'If (SmartTags("SDC\_TS_Nr") < SmartTags("DB_SDC_TS_IF_STATUS.HEADER.SEK_MIN")) Or (SmartTags("SDC\_TS_Nr") > SmartTags("DB_SDC_TS_IF_STATUS.HEADER.SEK_MAX")) Then
   '	If (SmartTags("SDC\_TS_Nr") < SmartTags("DB_SDC_TS_IF_STATUS_2.HEADER.SEK_MIN")) Or (SmartTags("SDC\_TS_Nr") > SmartTags("DB_SDC_TS_IF_STATUS_2.HEADER.SEK_MAX")) Then
   '		SmartTags("SDC\_TS_Nr") = 	SmartTags("DB_SDC_TS_IF_STATUS.HEADER.SEK_MIN")
   '	End If		
   'End If	
   	
   
   'If (SmartTags("SDC\_TS_Nr") < 1) Then
   '	SmartTags("SDC\_TS_Nr") = 1
   'End If	
   
   'TS_Nr = SmartTags("SDC\_TS_Nr")
   
   'If (SmartTags("SDC\_TS_Nr") >= SmartTags("DB_SDC_TS_IF_STATUS_2.HEADER.SEK_MIN")) And (SmartTags("SDC\_TS_Nr") <= SmartTags("DB_SDC_TS_IF_STATUS_2.HEADER.SEK_MAX")) Then
   '	SmartTags("_Byte_DB_SDC_TS_IF_STATUS.HEADER.DB_NR") = SmartTags("DB_SDC_TS_IF_STATUS_2.HEADER.DB_NR")	
   '	TS_Nr = SmartTags("SDC\_TS_Nr") - SmartTags("DB_SDC_TS_IF_STATUS_2.HEADER.SEK_MIN") + 1
   'End If	
   
   
   
   '##############################################
   ' VISU Sucht sich Sektions daten:
   '##############################################
   'Laenge_Data = SmartTags("DB_SDC_TS_IF_STATUS.HEADER.LAENGE_SEK_DATA")
   
   'Allg_Offset = SmartTags("DB_SDC_TS_IF_STATUS.HEADER.START_DAT")
   
   'OffsetTS = TS_Nr  * Laenge_Data - Laenge_Data + Allg_Offset
   
   'SmartTags("_Byte_DB_SDC_TS_IF_STATUS.SEK[XXX].VAL.EMS_ID") =						  0 + OffsetTS
   'SmartTags("_Byte_DB_SDC_TS_IF_STATUS.SEK[XXX].VAL.PROFIL") =						  2 + OffsetTS
   'SmartTags("_Byte_DB_SDC_TS_IF_STATUS.SEK[XXX].VAL.DRIVE_POS") =						  4 + OffsetTS
   'SmartTags("_Byte_DB_SDC_TS_IF_STATUS.SEK[XXX].VAL.HOIST_POS") =						  8 + OffsetTS
   'SmartTags("_Byte_DB_SDC_TS_IF_STATUS.SEK[XXX].VAL.TILT_POS") =						 10 + OffsetTS
   'SmartTags("_Byte_DB_SDC_TS_IF_STATUS.SEK[XXX].VAL.ERROR") =							 12 + OffsetTS
   'SmartTags("_Byte_DB_SDC_TS_IF_STATUS.SEK[XXX].VAL.DRIVE_POS_PERC") =				 14 + OffsetTS
   'SmartTags("_Byte_DB_SDC_TS_IF_STATUS.SEK[XXX].VAL.SEK") =							 16 + OffsetTS
   
   'SmartTags("_Byte_DB_SDC_TS_IF_STATUS.SEK[XXX].BIT1") =					 			 18 + OffsetTS
   'SmartTags("_Byte_DB_SDC_TS_IF_STATUS.SEK[XXX].BIT2") =					 			 20 + OffsetTS
   'SmartTags("_Byte_DB_SDC_TS_IF_STATUS.SEK[XXX].BIT3") =					 			 22 + OffsetTS
   'SmartTags("_Byte_DB_SDC_TS_IF_STATUS.SEK[XXX].BIT4") =					 			 24 + OffsetTS
   
   'SmartTags("_Byte_DB_SDC_TS_IF_STATUS.SEK[XXX].SORTE") =					 			 26 + OffsetTS
   
   'SmartTags("_Byte_DB_SDC_TS_IF_STATUS.SEK[XXX].FKT_SET") =				 			 30 + OffsetTS

VB script "SDC_TS_PARAMETER"
   'HINWEIS:
   ' Beim Erstellen von Skripten können Sie mit <Strg+Leertaste> vordefinierte 
   ' Systemfunktionen in das neue Skript einbinden.
   ' Das HMIRuntime-Objekt ermöglicht einfachen Zugriff auf die Objekte des
   ' WinCC flexible Objektmodells, ihre Methoden und ihre Eigenschaften.
   ' Für ein komfortables Auswählen einer Objektreferenz betätigen Sie bitte <Alt+Rechts>.
   ' Komplexe Skripte können Sie mit Sprachelementen der Programmiersprache
   ' VBScript erstellen.
   ' Der Zugriff auf WinCC flexible Variablen erfolgt direkt über den Variablennamen,
   ' z.B. Tag = 5
   
   '________________________________________________________________________________
   '
   
   ' Groiß Andreas
   ' Siemens AG Österreich 
   ' Linz Kraußstraße 1-7 
   ' RC-AT I-IA AS-FA-SO-AE2
   ' 01.08.2013
   
   Dim TS_Nr ' Sektion Number
   Dim TS_Profil_Nr ' Profil Number
   Dim Laenge_Data ' Länge TS Parameter
   Dim Laenge_Profil ' Länge TS Profil Parameter
   Dim Allg_Offset ' Allg Parameter Offset
   Dim Profil_Offset ' Allg Parameter Offset
   Dim HMISekDaten_Offset ' HMI Sektionsdaten Offset
   Dim HMI_Nr ' HMI Nummer
   
   ' INIT-------------------------------------------------------------
   SmartTags("SDC\DB_SDC_TS_PARAMETER\_TS_DB_Nr") = SmartTags("DB_SDC_TS_PARAMETER_HMI_HEADER.DB_NR")
   
   If (SmartTags("SDC\_TS_Nr") < SmartTags("DB_SDC_GLOBAL_SEK_MIN")) Or (SmartTags("SDC\_TS_Nr") > SmartTags("DB_SDC_GLOBAL_SEK_MAX")) Then
   	SmartTags("SDC\_TS_Nr") = 	SmartTags("DB_SDC_GLOBAL_SEK_MIN")
   End If	
   
   If (SmartTags("SDC\_TS_Nr") < 1) Then
   	SmartTags("SDC\_TS_Nr") = 1
   End If	
   
   'Anzahl Profile - 1 da 2 Profilparemter anmgezeigt werden
   If (SmartTags("SDC\DB_SDC_TS_PARAMETER\_TS_Profil_Nr") > (SmartTags("DB_SDC_TS_PARAMETER_1_HEADER.ANZ_PROFIL")- 1)) Or (SmartTags("SDC\DB_SDC_TS_PARAMETER\_TS_Profil_Nr") < 1 ) Then 
   	SmartTags("SDC\DB_SDC_TS_PARAMETER\_TS_Profil_Nr") = 1
   End If
   
   SmartTags("SDC\DB_SDC_TS_PARAMETER\_TS_Profil_Nr+1") = SmartTags("SDC\DB_SDC_TS_PARAMETER\_TS_Profil_Nr") + 1
   
   '##############################################
   ' S7 sucht sich Sektionsdaten:
   '##############################################
   
   	TS_Profil_Nr = SmartTags("SDC\DB_SDC_TS_PARAMETER\_TS_Profil_Nr")
   	
   	TS_Nr = SmartTags("SDC\_TS_Nr")
   	
   	Laenge_Data = SmartTags("DB_SDC_TS_PARAMETER_HMI_HEADER.LAENGE_SEK_DATA")
   	Laenge_Profil = SmartTags("DB_SDC_TS_PARAMETER_HMI_HEADER.LAENGE_PROFIL_DATA")
   	Allg_Offset = SmartTags("DB_SDC_TS_PARAMETER_HMI_HEADER.START_HMI")
   	Profil_Offset = SmartTags("DB_SDC_TS_PARAMETER_HMI_HEADER.OFFEST_PROFIL")
   	HMISekDaten_Offset = SmartTags("DB_SDC_TS_PARAMETER_HMI_HEADER.OFFEST_HMI_DATA")
   	HMI_Nr = SmartTags("_intern_Pult_Nr")